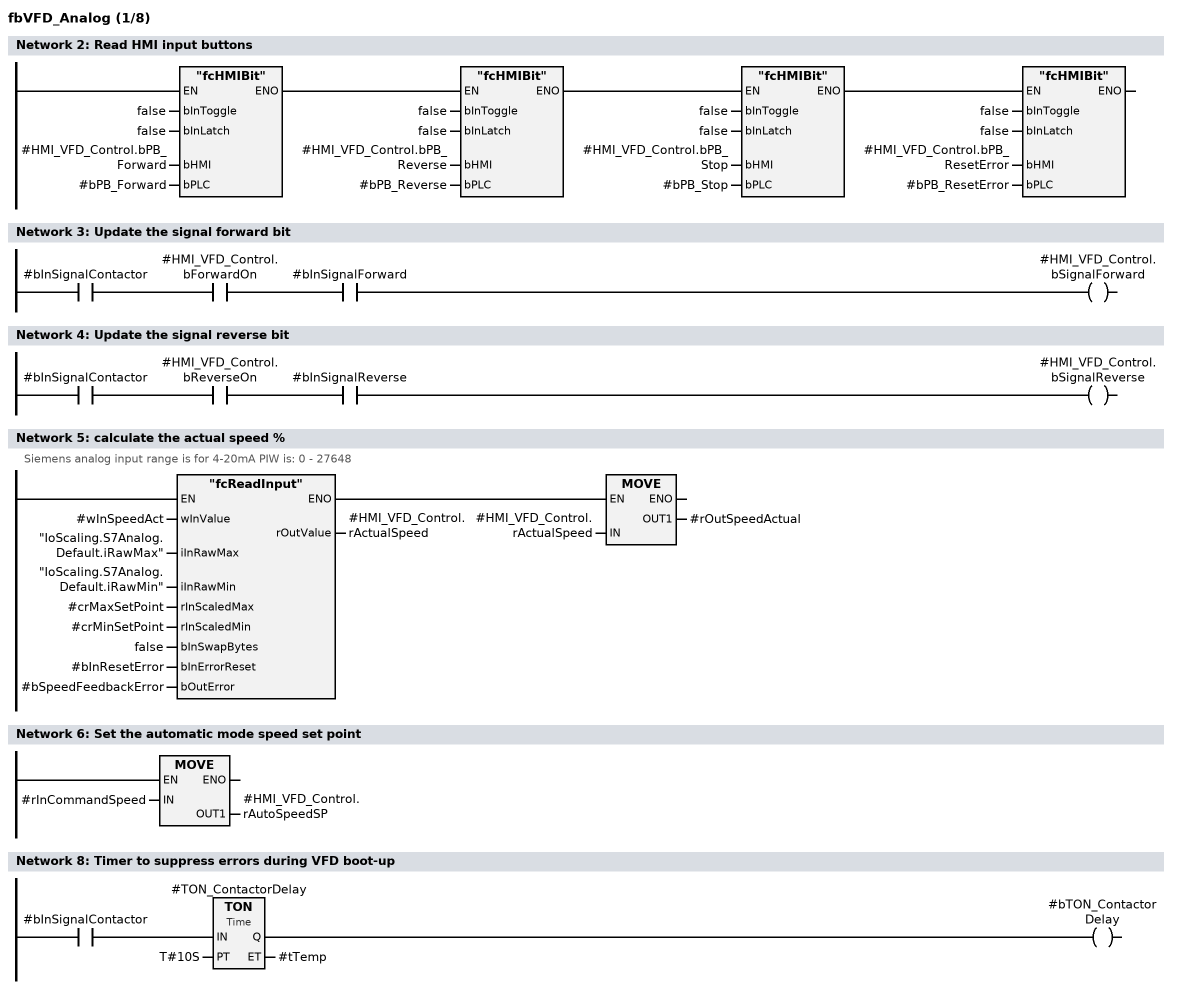
   RUNG wire#powerrail
      "fcHMIBit"(bInToggle := false, bInLatch := false, bHMI := #HMI_VFD_Control.bPB_Forward, bPLC := #bPB_Forward)
      "fcHMIBit"(bInToggle := false, bInLatch := false, bHMI := #HMI_VFD_Control.bPB_Reverse, bPLC := #bPB_Reverse)
      "fcHMIBit"(bInToggle := false, bInLatch := false, bHMI := #HMI_VFD_Control.bPB_Stop, bPLC := #bPB_Stop)
      "fcHMIBit"(bInToggle := false, bInLatch := false, bHMI := #HMI_VFD_Control.bPB_ResetError, bPLC := #bPB_ResetError)
   END_RUNG
   // the same network as SCL:
   "fcHMIBit"(bInToggle := false,
              bInLatch := false,
              bHMI := #HMI_VFD_Control.bPB_Forward,
              bPLC := #bPB_Forward,
              ENO => #_w1);
   "fcHMIBit"(EN := #_w1,
              bInToggle := false,
              bInLatch := false,
              bHMI := #HMI_VFD_Control.bPB_Reverse,
              bPLC := #bPB_Reverse,
              ENO => #_w2);
   "fcHMIBit"(EN := #_w2,
              bInToggle := false,
              bInLatch := false,
              bHMI := #HMI_VFD_Control.bPB_Stop,
              bPLC := #bPB_Stop,
              ENO => #_w3);
   IF #_w3 THEN
       "fcHMIBit"(bInToggle := false,
                  bInLatch := false,
                  bHMI := #HMI_VFD_Control.bPB_ResetError,
                  bPLC := #bPB_ResetError);
   END_IF;
END_REGION

REGION Network 3: Update the signal forward bit
   RUNG wire#powerrail
      Contact( #bInSignalContactor )
      Contact( #HMI_VFD_Control.bForwardOn )
      Contact( #bInSignalForward )
      Coil( #HMI_VFD_Control.bSignalForward )
   END_RUNG
   // the same network as SCL:
   #HMI_VFD_Control.bSignalForward := #bInSignalContactor AND #HMI_VFD_Control.bForwardOn AND #bInSignalForward;
END_REGION

REGION Network 4: Update the signal reverse bit
   RUNG wire#powerrail
      Contact( #bInSignalContactor )
      Contact( #HMI_VFD_Control.bReverseOn )
      Contact( #bInSignalReverse )
      Coil( #HMI_VFD_Control.bSignalReverse )
   END_RUNG
   // the same network as SCL:
   #HMI_VFD_Control.bSignalReverse := #bInSignalContactor AND #HMI_VFD_Control.bReverseOn AND #bInSignalReverse;
END_REGION

REGION Network 5: calculate the actual speed %
   // Siemens analog input range is for 4-20mA PIW is: 0 - 27648
   RUNG wire#powerrail
      "fcReadInput"(wInValue := #wInSpeedAct, iInRawMax := "IoScaling.S7Analog.Default.iRawMax", iInRawMin := "IoScaling.S7Analog.Default.iRawMin", rInScaledMax := #crMaxSetPoint, rInScaledMin := #crMinSetPoint, bInSwapBytes := false, bInErrorReset := #bInResetError, bOutError := #bSpeedFeedbackError, rOutValue => #HMI_VFD_Control.rActualSpeed)
      { S7_GenerateENO := "TRUE" } Move(in := #HMI_VFD_Control.rActualSpeed, out1 => #rOutSpeedActual)
   END_RUNG
   // the same network as SCL:
   "fcReadInput"(wInValue := #wInSpeedAct,
                 iInRawMax := "IoScaling.S7Analog.Default.iRawMax",
                 iInRawMin := "IoScaling.S7Analog.Default.iRawMin",
                 rInScaledMax := #crMaxSetPoint,
                 rInScaledMin := #crMinSetPoint,
                 bInSwapBytes := false,
                 bInErrorReset := #bInResetError,
                 bOutError := #bSpeedFeedbackError,
                 rOutValue => #HMI_VFD_Control.rActualSpeed,
                 ENO => #_w1);
   IF #_w1 THEN #rOutSpeedActual := #HMI_VFD_Control.rActualSpeed; END_IF;
END_REGION

REGION Network 6: Set the automatic mode speed set point
   RUNG wire#powerrail
      { S7_GenerateENO := "TRUE" } Move(in := #rInCommandSpeed, out1 => #HMI_VFD_Control.rAutoSpeedSP)
   END_RUNG
   // the same network as SCL:
   #HMI_VFD_Control.rAutoSpeedSP := #rInCommandSpeed;
END_REGION

REGION Network 7: --------------------------------------------------- Control Logic ------------------------------------------------------------
END_REGION

REGION Network 8: Timer to suppress errors during VFD boot-up
   #TON_ContactorDelay.TON(IN := #bInSignalContactor, PT := T#10S, ET => #tTemp);
   #bTON_ContactorDelay := #TON_ContactorDelay.Q;
END_REGION

REGION Network 9: Limit manual and auto set points to the max and min constants
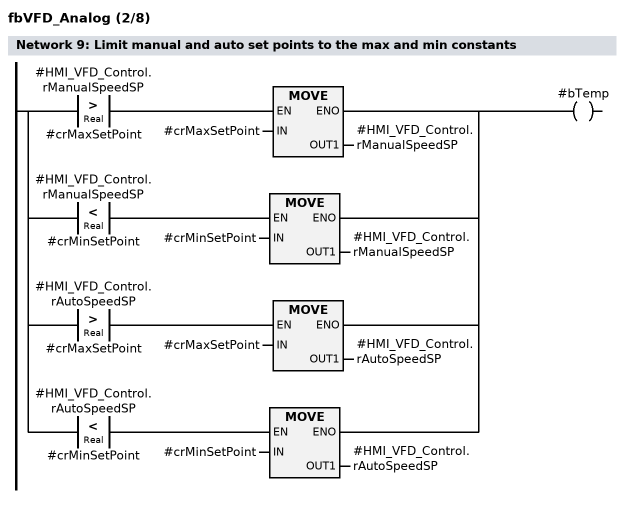
   RUNG wire#powerrail
      { S7_Templates := "SrcType := Real" } GT_Contact(in1 := #HMI_VFD_Control.rManualSpeedSP, in2 := #crMaxSetPoint)
      { S7_GenerateENO := "TRUE" } Move(in := #crMaxSetPoint, out1 => #HMI_VFD_Control.rManualSpeedSP)
      wire#w1
      Coil( #bTemp )
   END_RUNG
   RUNG wire#powerrail
      { S7_Templates := "SrcType := Real" } LT_Contact(in1 := #HMI_VFD_Control.rManualSpeedSP, in2 := #crMinSetPoint)
      { S7_GenerateENO := "TRUE" } Move(in := #crMinSetPoint, out1 => #HMI_VFD_Control.rManualSpeedSP)
   END_RUNG wire#w1
   RUNG wire#powerrail
      { S7_Templates := "SrcType := Real" } GT_Contact(in1 := #HMI_VFD_Control.rAutoSpeedSP, in2 := #crMaxSetPoint)
      { S7_GenerateENO := "TRUE" } Move(in := #crMaxSetPoint, out1 => #HMI_VFD_Control.rAutoSpeedSP)
   END_RUNG wire#w1
   RUNG wire#powerrail
      { S7_Templates := "SrcType := Real" } LT_Contact(in1 := #HMI_VFD_Control.rAutoSpeedSP, in2 := #crMinSetPoint)
      { S7_GenerateENO := "TRUE" } Move(in := #crMinSetPoint, out1 => #HMI_VFD_Control.rAutoSpeedSP)
   END_RUNG wire#w1
   // the same network as SCL:
   // ENO of a box is taken as its EN; it also drops when the box reports an error
   #_w1 := #HMI_VFD_Control.rManualSpeedSP > #crMaxSetPoint;
   IF #_w1 THEN #HMI_VFD_Control.rManualSpeedSP := #crMaxSetPoint; END_IF;
   #_w2 := #HMI_VFD_Control.rManualSpeedSP < #crMinSetPoint;
   IF #_w2 THEN #HMI_VFD_Control.rManualSpeedSP := #crMinSetPoint; END_IF;
   #_w3 := #HMI_VFD_Control.rAutoSpeedSP > #crMaxSetPoint;
   IF #_w3 THEN #HMI_VFD_Control.rAutoSpeedSP := #crMaxSetPoint; END_IF;
   #_w4 := #HMI_VFD_Control.rAutoSpeedSP < #crMinSetPoint;
   IF #_w4 THEN #HMI_VFD_Control.rAutoSpeedSP := #crMinSetPoint; END_IF;
   #bTemp := #_w1 OR #_w2 OR #_w3 OR #_w4;
END_REGION

REGION Network 10: Reset Errors
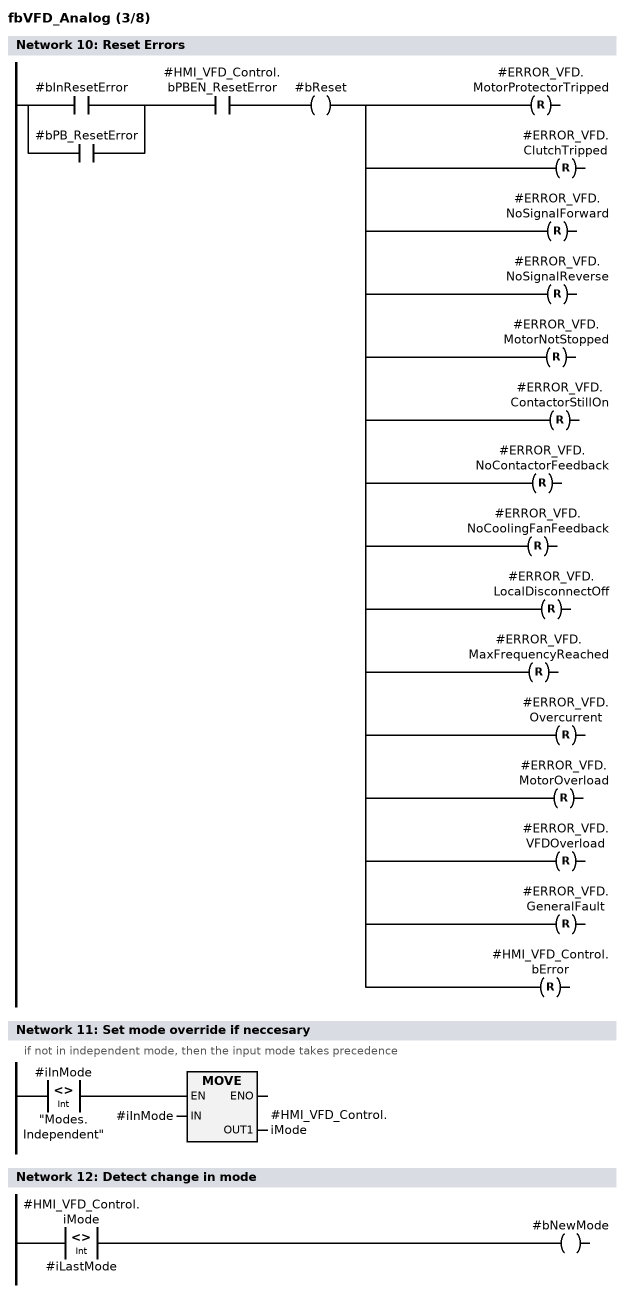
   RUNG wire#powerrail
      Contact( #bInResetError )
      wire#w1
      Contact( #HMI_VFD_Control.bPBEN_ResetError )
      Coil( #bReset )
      wire#w2
      R_Coil( #ERROR_VFD.MotorProtectorTripped )
   END_RUNG
   RUNG wire#powerrail
      Contact( #bPB_ResetError )
   END_RUNG wire#w1
   RUNG wire#w2
      R_Coil( #ERROR_VFD.ClutchTripped )
   END_RUNG
   RUNG wire#w2
      R_Coil( #ERROR_VFD.NoSignalForward )
   END_RUNG
   RUNG wire#w2
      R_Coil( #ERROR_VFD.NoSignalReverse )
   END_RUNG
   RUNG wire#w2
      R_Coil( #ERROR_VFD.MotorNotStopped )
   END_RUNG
   RUNG wire#w2
      R_Coil( #ERROR_VFD.ContactorStillOn )
   END_RUNG
   RUNG wire#w2
      R_Coil( #ERROR_VFD.NoContactorFeedback )
   END_RUNG
   RUNG wire#w2
      R_Coil( #ERROR_VFD.NoCoolingFanFeedback )
   END_RUNG
   RUNG wire#w2
      R_Coil( #ERROR_VFD.LocalDisconnectOff )
   END_RUNG
   RUNG wire#w2
      R_Coil( #ERROR_VFD.MaxFrequencyReached )
   END_RUNG
   RUNG wire#w2
      R_Coil( #ERROR_VFD.Overcurrent )
   END_RUNG
   RUNG wire#w2
      R_Coil( #ERROR_VFD.MotorOverload )
   END_RUNG
   RUNG wire#w2
      R_Coil( #ERROR_VFD.VFDOverload )
   END_RUNG
   RUNG wire#w2
      R_Coil( #ERROR_VFD.GeneralFault )
   END_RUNG
   RUNG wire#w2
      R_Coil( #HMI_VFD_Control.bError )
   END_RUNG
   // the same network as SCL:
   #bReset := (#bInResetError OR #bPB_ResetError) AND #HMI_VFD_Control.bPBEN_ResetError;
   IF #bReset THEN
       #ERROR_VFD.MotorProtectorTripped := FALSE;
       #ERROR_VFD.ClutchTripped := FALSE;
       #ERROR_VFD.NoSignalForward := FALSE;
       #ERROR_VFD.NoSignalReverse := FALSE;
       #ERROR_VFD.MotorNotStopped := FALSE;
       #ERROR_VFD.ContactorStillOn := FALSE;
       #ERROR_VFD.NoContactorFeedback := FALSE;
       #ERROR_VFD.NoCoolingFanFeedback := FALSE;
       #ERROR_VFD.LocalDisconnectOff := FALSE;
       #ERROR_VFD.MaxFrequencyReached := FALSE;
       #ERROR_VFD.Overcurrent := FALSE;
       #ERROR_VFD.MotorOverload := FALSE;
       #ERROR_VFD.VFDOverload := FALSE;
       #ERROR_VFD.GeneralFault := FALSE;
       #HMI_VFD_Control.bError := FALSE;
   END_IF;
END_REGION

REGION Network 11: Set mode override if neccesary
   // if not in independent mode, then the input mode takes precedence
   RUNG wire#powerrail
      { S7_Templates := "SrcType := Int" } NE_Contact(in1 := #iInMode, in2 := "Modes.Independent")
      { S7_GenerateENO := "TRUE" } Move(in := #iInMode, out1 => #HMI_VFD_Control.iMode)
   END_RUNG
   // the same network as SCL:
   IF #iInMode <> "Modes.Independent" THEN #HMI_VFD_Control.iMode := #iInMode; END_IF;
END_REGION

REGION Network 12: Detect change in mode
   RUNG wire#powerrail
      { S7_Templates := "SrcType := Int" } NE_Contact(in1 := #HMI_VFD_Control.iMode, in2 := #iLastMode)
      Coil( #bNewMode )
   END_RUNG
   // the same network as SCL:
   #bNewMode := #HMI_VFD_Control.iMode <> #iLastMode;
END_REGION

REGION Network 13: Keep track of last mode
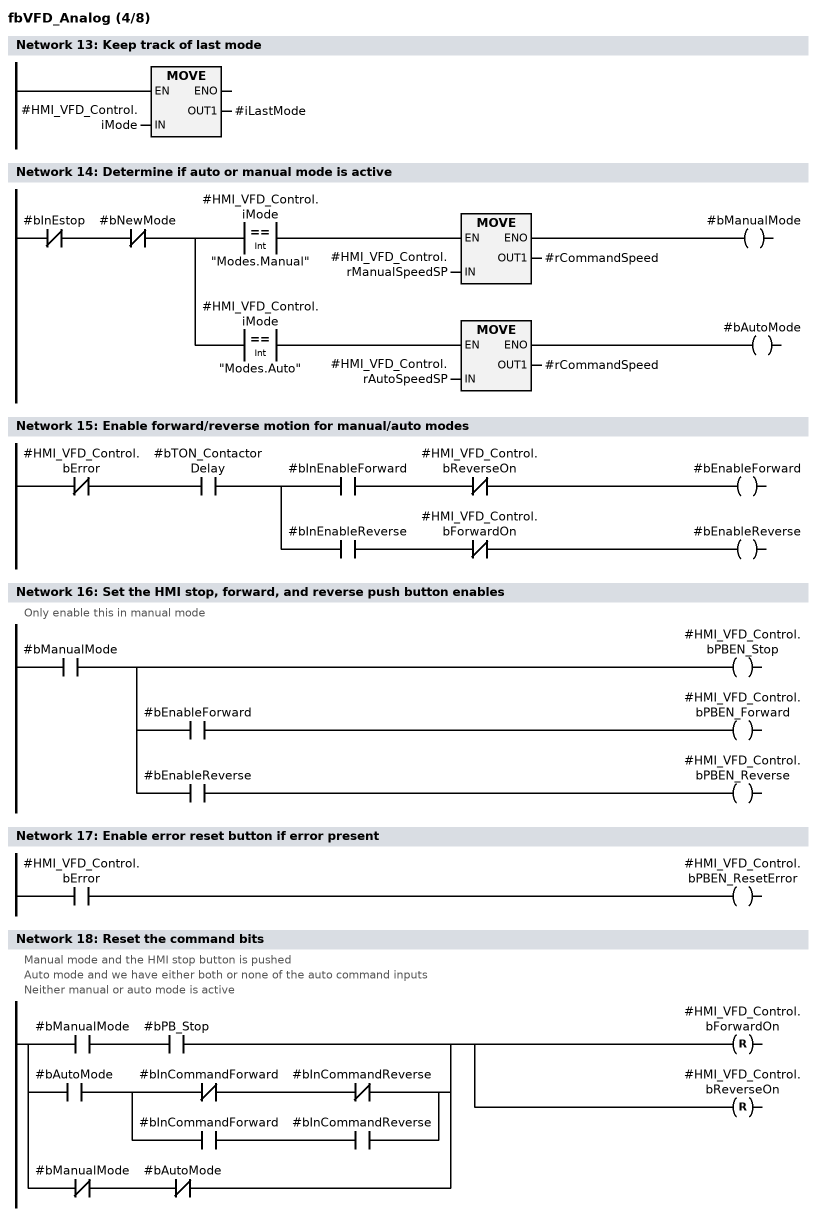
   RUNG wire#powerrail
      { S7_GenerateENO := "TRUE" } Move(in := #HMI_VFD_Control.iMode, out1 => #iLastMode)
   END_RUNG
   // the same network as SCL:
   #iLastMode := #HMI_VFD_Control.iMode;
END_REGION

REGION Network 14: Determine if auto or manual mode is active
   RUNG wire#powerrail
      I_Contact( #bInEstop )
      I_Contact( #bNewMode )
      wire#w1
      { S7_Templates := "SrcType := Int" } EQ_Contact(in1 := #HMI_VFD_Control.iMode, in2 := "Modes.Manual")
      { S7_GenerateENO := "TRUE" } Move(in := #HMI_VFD_Control.rManualSpeedSP, out1 => #rCommandSpeed)
      Coil( #bManualMode )
   END_RUNG
   RUNG wire#w1
      { S7_Templates := "SrcType := Int" } EQ_Contact(in1 := #HMI_VFD_Control.iMode, in2 := "Modes.Auto")
      { S7_GenerateENO := "TRUE" } Move(in := #HMI_VFD_Control.rAutoSpeedSP, out1 => #rCommandSpeed)
      Coil( #bAutoMode )
   END_RUNG
   // the same network as SCL:
   // ENO of a box is taken as its EN; it also drops when the box reports an error
   #_w1 := NOT #bInEstop AND NOT #bNewMode;
   #_w2 := #_w1 AND (#HMI_VFD_Control.iMode = "Modes.Manual");
   IF #_w2 THEN #rCommandSpeed := #HMI_VFD_Control.rManualSpeedSP; END_IF;
   #bManualMode := #_w2;
   #_w3 := #_w1 AND (#HMI_VFD_Control.iMode = "Modes.Auto");
   IF #_w3 THEN #rCommandSpeed := #HMI_VFD_Control.rAutoSpeedSP; END_IF;
   #bAutoMode := #_w3;
END_REGION

REGION Network 15: Enable forward/reverse motion for manual/auto modes
   RUNG wire#powerrail
      I_Contact( #HMI_VFD_Control.bError )
      Contact( #bTON_ContactorDelay )
      wire#w1
      Contact( #bInEnableForward )
      I_Contact( #HMI_VFD_Control.bReverseOn )
      Coil( #bEnableForward )
   END_RUNG
   RUNG wire#w1
      Contact( #bInEnableReverse )
      I_Contact( #HMI_VFD_Control.bForwardOn )
      Coil( #bEnableReverse )
   END_RUNG
   // the same network as SCL:
   #_w1 := NOT #HMI_VFD_Control.bError AND #bTON_ContactorDelay;
   #bEnableForward := #_w1 AND #bInEnableForward AND NOT #HMI_VFD_Control.bReverseOn;
   #bEnableReverse := #_w1 AND #bInEnableReverse AND NOT #HMI_VFD_Control.bForwardOn;
END_REGION

REGION Network 16: Set the HMI stop, forward, and reverse push button enables
   // Only enable this in manual mode
   RUNG wire#powerrail
      Contact( #bManualMode )
      wire#w1
      Coil( #HMI_VFD_Control.bPBEN_Stop )
   END_RUNG
   RUNG wire#w1
      Contact( #bEnableForward )
      Coil( #HMI_VFD_Control.bPBEN_Forward )
   END_RUNG
   RUNG wire#w1
      Contact( #bEnableReverse )
      Coil( #HMI_VFD_Control.bPBEN_Reverse )
   END_RUNG
   // the same network as SCL:
   #HMI_VFD_Control.bPBEN_Stop := #bManualMode;
   #HMI_VFD_Control.bPBEN_Forward := #bManualMode AND #bEnableForward;
   #HMI_VFD_Control.bPBEN_Reverse := #bManualMode AND #bEnableReverse;
END_REGION

REGION Network 17: Enable error reset button if error present
   RUNG wire#powerrail
      Contact( #HMI_VFD_Control.bError )
      Coil( #HMI_VFD_Control.bPBEN_ResetError )
   END_RUNG
   // the same network as SCL:
   #HMI_VFD_Control.bPBEN_ResetError := #HMI_VFD_Control.bError;
END_REGION

REGION Network 18: Reset the command bits
   // Manual mode and the HMI stop button is pushed
   // Auto mode and we have either both or none of the auto command inputs
   // Neither manual or auto mode is active
   RUNG wire#powerrail
      Contact( #bManualMode )
      Contact( #bPB_Stop )
      wire#w1
      R_Coil( #HMI_VFD_Control.bForwardOn )
   END_RUNG
   RUNG wire#powerrail
      Contact( #bAutoMode )
      wire#w2
      I_Contact( #bInCommandForward )
      I_Contact( #bInCommandReverse )
   END_RUNG wire#w1
   RUNG wire#w2
      Contact( #bInCommandForward )
      Contact( #bInCommandReverse )
   END_RUNG wire#w1
   RUNG wire#powerrail
      I_Contact( #bManualMode )
      I_Contact( #bAutoMode )
   END_RUNG wire#w1
   RUNG wire#w1
      R_Coil( #HMI_VFD_Control.bReverseOn )
   END_RUNG
   // the same network as SCL:
   IF (#bManualMode AND #bPB_Stop) OR (#bAutoMode AND ((NOT #bInCommandForward AND NOT #bInCommandReverse) OR (#bInCommandForward AND #bInCommandReverse))) OR (NOT #bManualMode AND NOT #bAutoMode) THEN
       #HMI_VFD_Control.bForwardOn := FALSE;
       #HMI_VFD_Control.bReverseOn := FALSE;
   END_IF;
END_REGION

REGION Network 19: Start forward request
   // Manual mode and only a start forward button is pressed and enabled
   // Auto mode when we receive a auto command and it is enabled
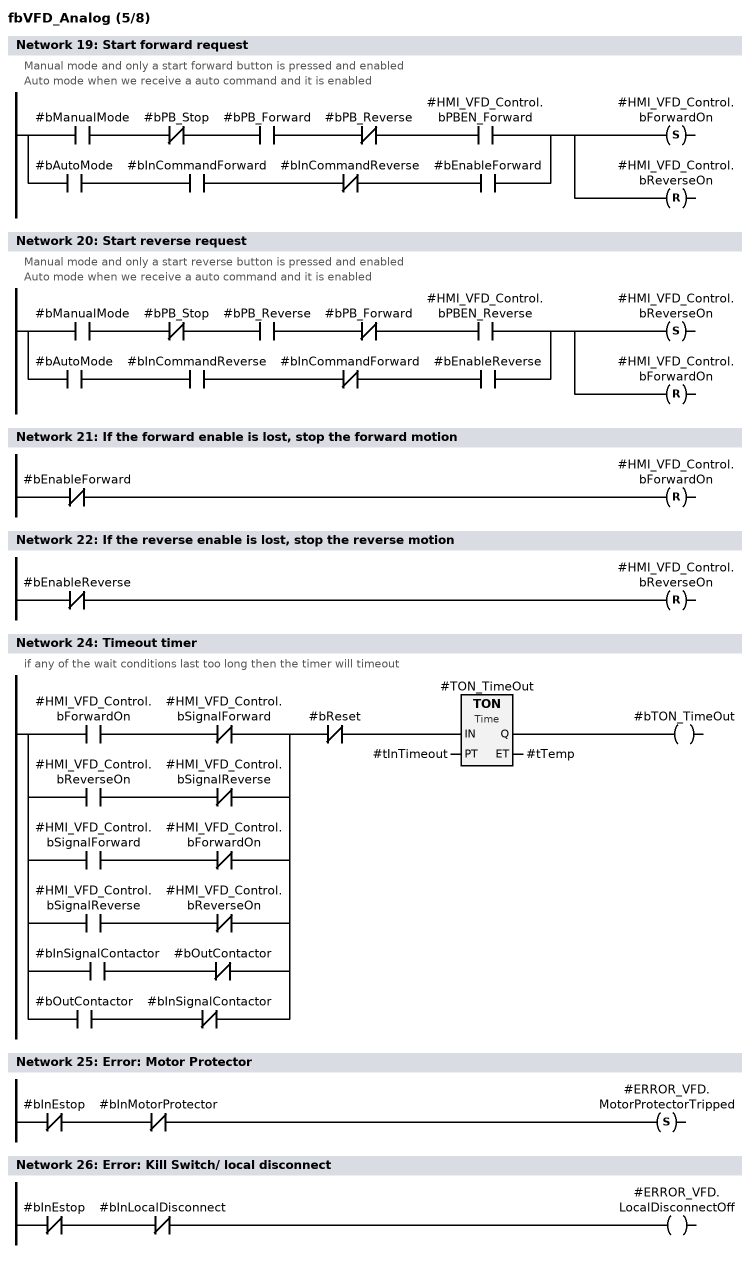
   RUNG wire#powerrail
      Contact( #bManualMode )
      I_Contact( #bPB_Stop )
      Contact( #bPB_Forward )
      I_Contact( #bPB_Reverse )
      Contact( #HMI_VFD_Control.bPBEN_Forward )
      wire#w1
      S_Coil( #HMI_VFD_Control.bForwardOn )
   END_RUNG
   RUNG wire#powerrail
      Contact( #bAutoMode )
      Contact( #bInCommandForward )
      I_Contact( #bInCommandReverse )
      Contact( #bEnableForward )
   END_RUNG wire#w1
   RUNG wire#w1
      R_Coil( #HMI_VFD_Control.bReverseOn )
   END_RUNG
   // the same network as SCL:
   IF (#bManualMode AND NOT #bPB_Stop AND #bPB_Forward AND NOT #bPB_Reverse AND #HMI_VFD_Control.bPBEN_Forward) OR (#bAutoMode AND #bInCommandForward AND NOT #bInCommandReverse AND #bEnableForward) THEN
       #HMI_VFD_Control.bForwardOn := TRUE;
       #HMI_VFD_Control.bReverseOn := FALSE;
   END_IF;
END_REGION

REGION Network 20: Start reverse request
   // Manual mode and only a start reverse button is pressed and enabled
   // Auto mode when we receive a auto command and it is enabled
   RUNG wire#powerrail
      Contact( #bManualMode )
      I_Contact( #bPB_Stop )
      Contact( #bPB_Reverse )
      I_Contact( #bPB_Forward )
      Contact( #HMI_VFD_Control.bPBEN_Reverse )
      wire#w1
      S_Coil( #HMI_VFD_Control.bReverseOn )
   END_RUNG
   RUNG wire#powerrail
      Contact( #bAutoMode )
      Contact( #bInCommandReverse )
      I_Contact( #bInCommandForward )
      Contact( #bEnableReverse )
   END_RUNG wire#w1
   RUNG wire#w1
      R_Coil( #HMI_VFD_Control.bForwardOn )
   END_RUNG
   // the same network as SCL:
   IF (#bManualMode AND NOT #bPB_Stop AND #bPB_Reverse AND NOT #bPB_Forward AND #HMI_VFD_Control.bPBEN_Reverse) OR (#bAutoMode AND #bInCommandReverse AND NOT #bInCommandForward AND #bEnableReverse) THEN
       #HMI_VFD_Control.bReverseOn := TRUE;
       #HMI_VFD_Control.bForwardOn := FALSE;
   END_IF;
END_REGION

REGION Network 21: If the forward enable is lost, stop the forward motion
   RUNG wire#powerrail
      I_Contact( #bEnableForward )
      R_Coil( #HMI_VFD_Control.bForwardOn )
   END_RUNG
   // the same network as SCL:
   IF NOT #bEnableForward THEN #HMI_VFD_Control.bForwardOn := FALSE; END_IF;
END_REGION

REGION Network 22: If the reverse enable is lost, stop the reverse motion
   RUNG wire#powerrail
      I_Contact( #bEnableReverse )
      R_Coil( #HMI_VFD_Control.bReverseOn )
   END_RUNG
   // the same network as SCL:
   IF NOT #bEnableReverse THEN #HMI_VFD_Control.bReverseOn := FALSE; END_IF;
END_REGION

REGION Network 23: --------------------------------------------------------- Errors ------------------------------------------------------------------
END_REGION

REGION Network 24: Timeout timer
   // if any of the wait conditions last too long then the timer will timeout
   #TON_TimeOut.TON(IN := ((#HMI_VFD_Control.bForwardOn AND NOT #HMI_VFD_Control.bSignalForward) OR (#HMI_VFD_Control.bReverseOn AND NOT #HMI_VFD_Control.bSignalReverse) OR (#HMI_VFD_Control.bSignalForward AND NOT #HMI_VFD_Control.bForwardOn) OR (#HMI_VFD_Control.bSignalReverse AND NOT #HMI_VFD_Control.bReverseOn) OR (#bInSignalContactor AND NOT #bOutContactor) OR (#bOutContactor AND NOT #bInSignalContactor)) AND NOT #bReset,
                    PT := #tInTimeout,
                    ET => #tTemp);
   #bTON_TimeOut := #TON_TimeOut.Q;
END_REGION

REGION Network 25: Error: Motor Protector
   RUNG wire#powerrail
      I_Contact( #bInEstop )
      I_Contact( #bInMotorProtector )
      S_Coil( #ERROR_VFD.MotorProtectorTripped )
   END_RUNG
   // the same network as SCL:
   IF NOT #bInEstop AND NOT #bInMotorProtector THEN #ERROR_VFD.MotorProtectorTripped := TRUE; END_IF;
END_REGION

REGION Network 26: Error: Kill Switch/ local disconnect
   RUNG wire#powerrail
      I_Contact( #bInEstop )
      I_Contact( #bInLocalDisconnect )
      Coil( #ERROR_VFD.LocalDisconnectOff )
   END_RUNG
   // the same network as SCL:
   #ERROR_VFD.LocalDisconnectOff := NOT #bInEstop AND NOT #bInLocalDisconnect;
END_REGION

REGION Network 27: Error Clutch
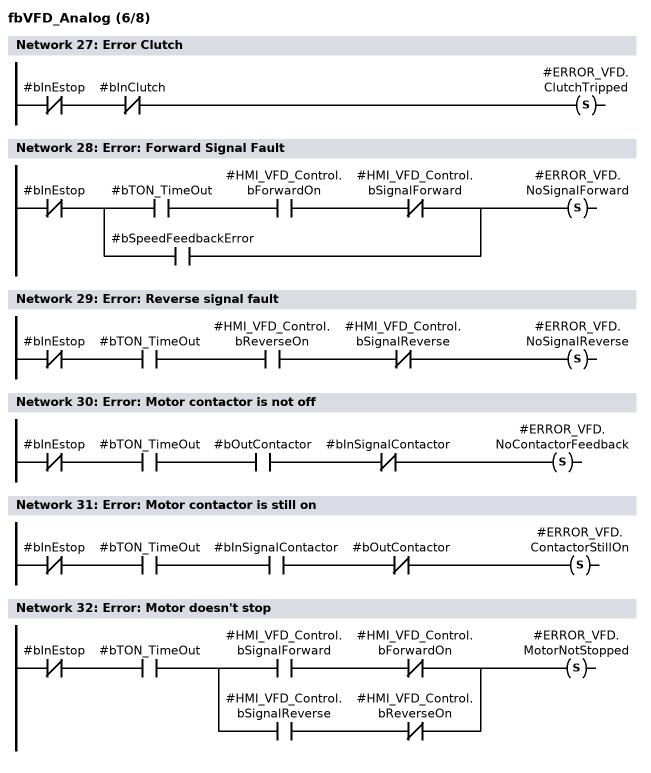
   RUNG wire#powerrail
      I_Contact( #bInEstop )
      I_Contact( #bInClutch )
      S_Coil( #ERROR_VFD.ClutchTripped )
   END_RUNG
   // the same network as SCL:
   IF NOT #bInEstop AND NOT #bInClutch THEN #ERROR_VFD.ClutchTripped := TRUE; END_IF;
END_REGION

REGION Network 28: Error: Forward Signal Fault
   RUNG wire#powerrail
      I_Contact( #bInEstop )
      wire#w1
      Contact( #bTON_TimeOut )
      Contact( #HMI_VFD_Control.bForwardOn )
      I_Contact( #HMI_VFD_Control.bSignalForward )
      wire#w2
      S_Coil( #ERROR_VFD.NoSignalForward )
   END_RUNG
   RUNG wire#w1
      Contact( #bSpeedFeedbackError )
   END_RUNG wire#w2
   // the same network as SCL:
   IF NOT #bInEstop AND ((#bTON_TimeOut AND #HMI_VFD_Control.bForwardOn AND NOT #HMI_VFD_Control.bSignalForward) OR #bSpeedFeedbackError) THEN
       #ERROR_VFD.NoSignalForward := TRUE;
   END_IF;
END_REGION

REGION Network 29: Error: Reverse signal fault
   RUNG wire#powerrail
      I_Contact( #bInEstop )
      Contact( #bTON_TimeOut )
      Contact( #HMI_VFD_Control.bReverseOn )
      I_Contact( #HMI_VFD_Control.bSignalReverse )
      S_Coil( #ERROR_VFD.NoSignalReverse )
   END_RUNG
   // the same network as SCL:
   IF NOT #bInEstop AND #bTON_TimeOut AND #HMI_VFD_Control.bReverseOn AND NOT #HMI_VFD_Control.bSignalReverse THEN
       #ERROR_VFD.NoSignalReverse := TRUE;
   END_IF;
END_REGION

REGION Network 30: Error: Motor contactor is not off
   RUNG wire#powerrail
      I_Contact( #bInEstop )
      Contact( #bTON_TimeOut )
      Contact( #bOutContactor )
      I_Contact( #bInSignalContactor )
      S_Coil( #ERROR_VFD.NoContactorFeedback )
   END_RUNG
   // the same network as SCL:
   IF NOT #bInEstop AND #bTON_TimeOut AND #bOutContactor AND NOT #bInSignalContactor THEN
       #ERROR_VFD.NoContactorFeedback := TRUE;
   END_IF;
END_REGION

REGION Network 31: Error: Motor contactor is still on
   RUNG wire#powerrail
      I_Contact( #bInEstop )
      Contact( #bTON_TimeOut )
      Contact( #bInSignalContactor )
      I_Contact( #bOutContactor )
      S_Coil( #ERROR_VFD.ContactorStillOn )
   END_RUNG
   // the same network as SCL:
   IF NOT #bInEstop AND #bTON_TimeOut AND #bInSignalContactor AND NOT #bOutContactor THEN
       #ERROR_VFD.ContactorStillOn := TRUE;
   END_IF;
END_REGION

REGION Network 32: Error: Motor doesn't stop
   RUNG wire#powerrail
      I_Contact( #bInEstop )
      Contact( #bTON_TimeOut )
      wire#w1
      Contact( #HMI_VFD_Control.bSignalForward )
      I_Contact( #HMI_VFD_Control.bForwardOn )
      wire#w2
      S_Coil( #ERROR_VFD.MotorNotStopped )
   END_RUNG
   RUNG wire#w1
      Contact( #HMI_VFD_Control.bSignalReverse )
      I_Contact( #HMI_VFD_Control.bReverseOn )
   END_RUNG wire#w2
   // the same network as SCL:
   IF NOT #bInEstop AND #bTON_TimeOut AND ((#HMI_VFD_Control.bSignalForward AND NOT #HMI_VFD_Control.bForwardOn) OR (#HMI_VFD_Control.bSignalReverse AND NOT #HMI_VFD_Control.bReverseOn)) THEN
       #ERROR_VFD.MotorNotStopped := TRUE;
   END_IF;
END_REGION

REGION Network 33: Scroll errors on the HMI
   // This block loops through all of the possible errors and displays them on the HMI 
   // by setting an index value for each error bit.
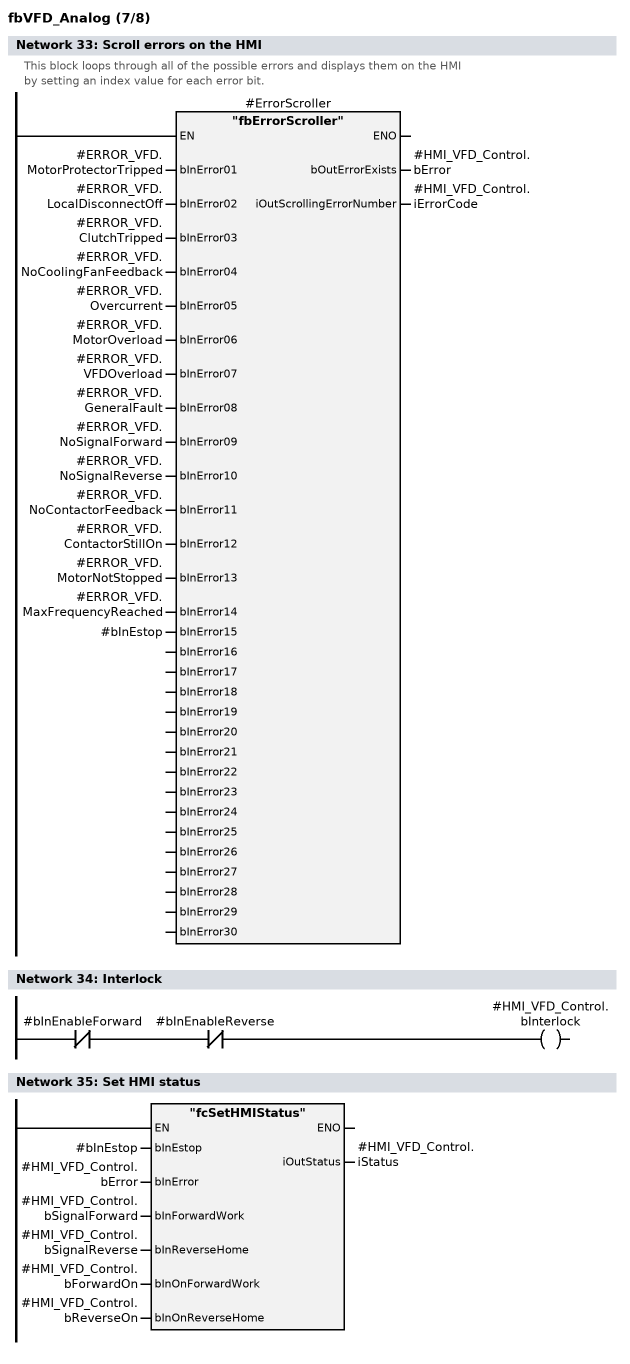
   RUNG wire#powerrail
      #ErrorScroller(bInError01 := #ERROR_VFD.MotorProtectorTripped, bInError02 := #ERROR_VFD.LocalDisconnectOff, bInError03 := #ERROR_VFD.ClutchTripped, bInError04 := #ERROR_VFD.NoCoolingFanFeedback, bInError05 := #ERROR_VFD.Overcurrent, bInError06 := #ERROR_VFD.MotorOverload, bInError07 := #ERROR_VFD.VFDOverload, bInError08 := #ERROR_VFD.GeneralFault, bInError09 := #ERROR_VFD.NoSignalForward, bInError10 := #ERROR_VFD.NoSignalReverse, bInError11 := #ERROR_VFD.NoContactorFeedback, bInError12 := #ERROR_VFD.ContactorStillOn, bInError13 := #ERROR_VFD.MotorNotStopped, bInError14 := #ERROR_VFD.MaxFrequencyReached, bInError15 := #bInEstop, bInError16 :=, bInError17 :=, bInError18 :=, bInError19 :=, bInError20 :=, bInError21 :=, bInError22 :=, bInError23 :=, bInError24 :=, bInError25 :=, bInError26 :=, bInError27 :=, bInError28 :=, bInError29 :=, bInError30 :=, bOutErrorExists => #HMI_VFD_Control.bError, iOutScrollingErrorNumber => #HMI_VFD_Control.iErrorCode)
   END_RUNG
   // the same network as SCL:
   #ErrorScroller(bInError01 := #ERROR_VFD.MotorProtectorTripped,   // "fbErrorScroller"
                  bInError02 := #ERROR_VFD.LocalDisconnectOff,
                  bInError03 := #ERROR_VFD.ClutchTripped,
                  bInError04 := #ERROR_VFD.NoCoolingFanFeedback,
                  bInError05 := #ERROR_VFD.Overcurrent,
                  bInError06 := #ERROR_VFD.MotorOverload,
                  bInError07 := #ERROR_VFD.VFDOverload,
                  bInError08 := #ERROR_VFD.GeneralFault,
                  bInError09 := #ERROR_VFD.NoSignalForward,
                  bInError10 := #ERROR_VFD.NoSignalReverse,
                  bInError11 := #ERROR_VFD.NoContactorFeedback,
                  bInError12 := #ERROR_VFD.ContactorStillOn,
                  bInError13 := #ERROR_VFD.MotorNotStopped,
                  bInError14 := #ERROR_VFD.MaxFrequencyReached,
                  bInError15 := #bInEstop,
                  bOutErrorExists => #HMI_VFD_Control.bError,
                  iOutScrollingErrorNumber => #HMI_VFD_Control.iErrorCode);
END_REGION

REGION Network 34: Interlock
   RUNG wire#powerrail
      I_Contact( #bInEnableForward )
      I_Contact( #bInEnableReverse )
      Coil( #HMI_VFD_Control.bInterlock )
   END_RUNG
   // the same network as SCL:
   #HMI_VFD_Control.bInterlock := NOT #bInEnableForward AND NOT #bInEnableReverse;
END_REGION

REGION Network 35: Set HMI status
   RUNG wire#powerrail
      "fcSetHMIStatus"(bInEstop := #bInEstop, bInError := #HMI_VFD_Control.bError, bInForwardWork := #HMI_VFD_Control.bSignalForward, bInReverseHome := #HMI_VFD_Control.bSignalReverse, bInOnForwardWork := #HMI_VFD_Control.bForwardOn, bInOnReverseHome := #HMI_VFD_Control.bReverseOn, iOutStatus => #HMI_VFD_Control.iStatus)
   END_RUNG
   // the same network as SCL:
   "fcSetHMIStatus"(bInEstop := #bInEstop,
                    bInError := #HMI_VFD_Control.bError,
                    bInForwardWork := #HMI_VFD_Control.bSignalForward,
                    bInReverseHome := #HMI_VFD_Control.bSignalReverse,
                    bInOnForwardWork := #HMI_VFD_Control.bForwardOn,
                    bInOnReverseHome := #HMI_VFD_Control.bReverseOn,
                    iOutStatus => #HMI_VFD_Control.iStatus);
END_REGION

REGION Network 36: -------------------------------------------------------- Outputs -------------------------------------------------------
END_REGION

REGION Network 37: Output: Forward
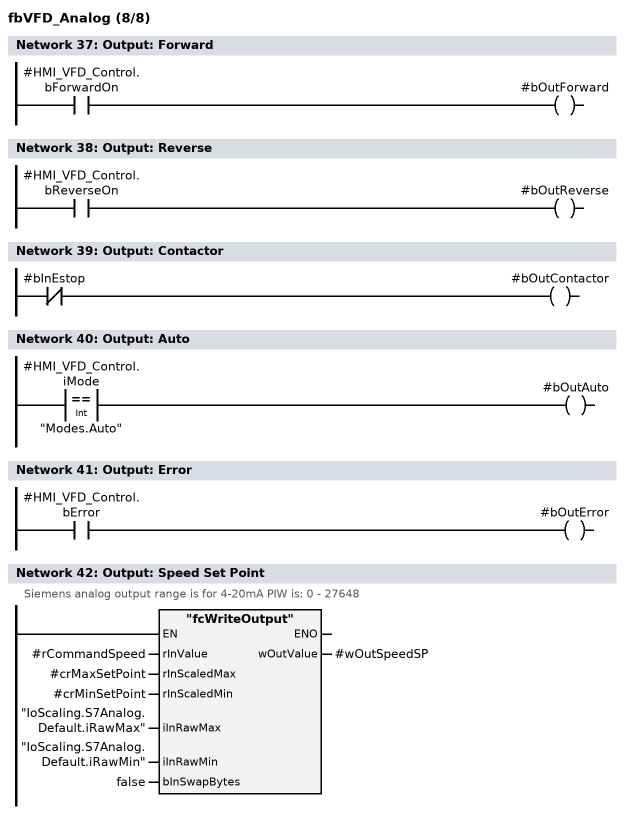
   RUNG wire#powerrail
      Contact( #HMI_VFD_Control.bForwardOn )
      Coil( #bOutForward )
   END_RUNG
   // the same network as SCL:
   #bOutForward := #HMI_VFD_Control.bForwardOn;
END_REGION

REGION Network 38: Output: Reverse
   RUNG wire#powerrail
      Contact( #HMI_VFD_Control.bReverseOn )
      Coil( #bOutReverse )
   END_RUNG
   // the same network as SCL:
   #bOutReverse := #HMI_VFD_Control.bReverseOn;
END_REGION

REGION Network 39: Output: Contactor
   RUNG wire#powerrail
      I_Contact( #bInEstop )
      Coil( #bOutContactor )
   END_RUNG
   // the same network as SCL:
   #bOutContactor := NOT #bInEstop;
END_REGION

REGION Network 40: Output: Auto
   RUNG wire#powerrail
      { S7_Templates := "SrcType := Int" } EQ_Contact(in1 := #HMI_VFD_Control.iMode, in2 := "Modes.Auto")
      Coil( #bOutAuto )
   END_RUNG
   // the same network as SCL:
   #bOutAuto := #HMI_VFD_Control.iMode = "Modes.Auto";
END_REGION

REGION Network 41: Output: Error
   RUNG wire#powerrail
      Contact( #HMI_VFD_Control.bError )
      Coil( #bOutError )
   END_RUNG
   // the same network as SCL:
   #bOutError := #HMI_VFD_Control.bError;
END_REGION

REGION Network 42: Output: Speed Set Point
   // Siemens analog output range is for 4-20mA PIW is: 0 - 27648
   RUNG wire#powerrail
      "fcWriteOutput"(rInValue := #rCommandSpeed, rInScaledMax := #crMaxSetPoint, rInScaledMin := #crMinSetPoint, iInRawMax := "IoScaling.S7Analog.Default.iRawMax", iInRawMin := "IoScaling.S7Analog.Default.iRawMin", bInSwapBytes := false, wOutValue => #wOutSpeedSP)
   END_RUNG
   // the same network as SCL:
   "fcWriteOutput"(rInValue := #rCommandSpeed,
                   rInScaledMax := #crMaxSetPoint,
                   rInScaledMin := #crMinSetPoint,
                   iInRawMax := "IoScaling.S7Analog.Default.iRawMax",
                   iInRawMin := "IoScaling.S7Analog.Default.iRawMin",
                   bInSwapBytes := false,
                   wOutValue => #wOutSpeedSP);
END_REGION
END_FUNCTION_BLOCK

FUNCTION_BLOCK "fbMotor_Reversing"   // FB130, LAD
TITLE = Controls a reversing motor contactor
{ S7_Optimized_Access := 'FALSE' }
VERSION : 0.1
   VAR_TEMP   // added for the SCL form of the ladder/FBD networks
      _w1 : Bool;
      _w2 : Bool;
      _w3 : Bool;
   END_VAR
BEGIN

REGION Network 1: --------------------------------------------------------- Inputs ------------------------------------------------------------------
END_REGION

REGION Network 2: Read HMI input buttons